REGION Network 8: FT-2011: R-201 Tank Flow from T-101 Totalizer
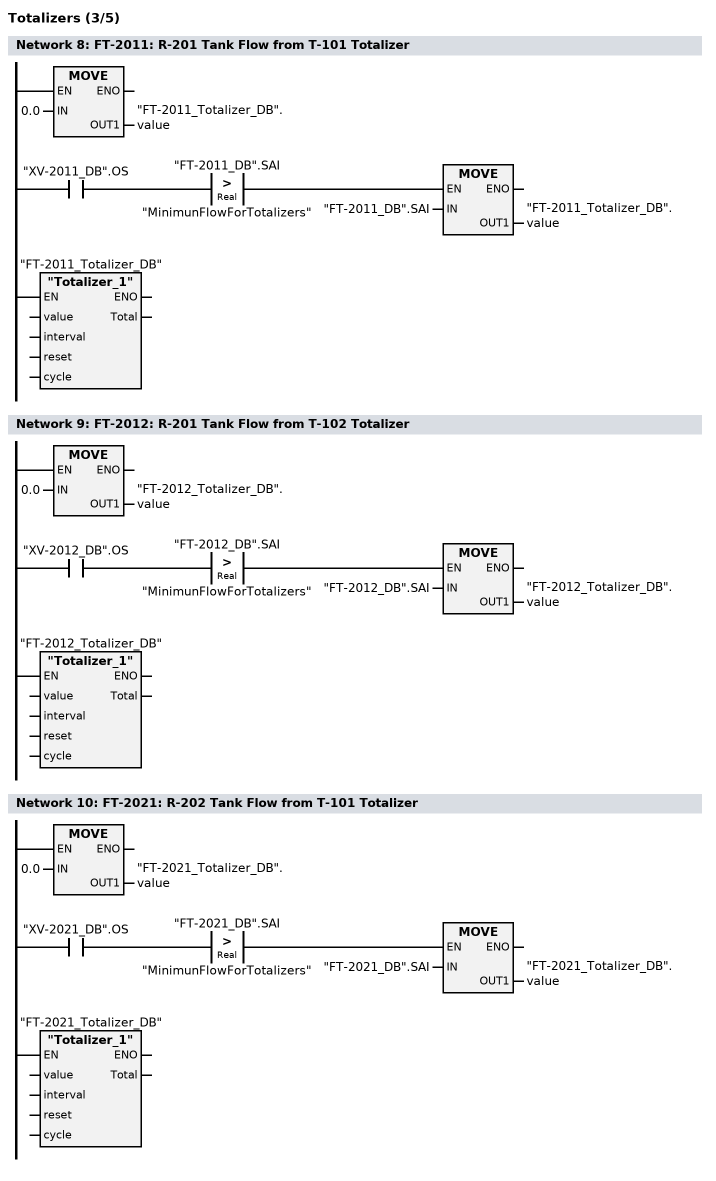
   RUNG wire#powerrail
      { S7_GenerateENO := "TRUE" } Move(in := 0.0, out1 => "FT-2011_Totalizer_DB".value)
   END_RUNG
   RUNG wire#powerrail
      Contact( "XV-2011_DB".OS )
      { S7_Templates := "SrcType := Real" } GT_Contact(in1 := "FT-2011_DB".SAI, in2 := "MinimunFlowForTotalizers")
      { S7_GenerateENO := "TRUE" } Move(in := "FT-2011_DB".SAI, out1 => "FT-2011_Totalizer_DB".value)
   END_RUNG
   RUNG wire#powerrail
      "FT-2011_Totalizer_DB"(value :=, interval :=, reset :=, cycle :=, Total =>)
   END_RUNG
   // the same network as SCL:
   "FT-2011_Totalizer_DB".value := 0.0;
   IF "XV-2011_DB".OS AND ("FT-2011_DB".SAI > "MinimunFlowForTotalizers") THEN
       "FT-2011_Totalizer_DB".value := "FT-2011_DB".SAI;
   END_IF;
   "FT-2011_Totalizer_DB"();   // "Totalizer_1"
END_REGION

REGION Network 9: FT-2012: R-201 Tank Flow from T-102 Totalizer
   RUNG wire#powerrail
      { S7_GenerateENO := "TRUE" } Move(in := 0.0, out1 => "FT-2012_Totalizer_DB".value)
   END_RUNG
   RUNG wire#powerrail
      Contact( "XV-2012_DB".OS )
      { S7_Templates := "SrcType := Real" } GT_Contact(in1 := "FT-2012_DB".SAI, in2 := "MinimunFlowForTotalizers")
      { S7_GenerateENO := "TRUE" } Move(in := "FT-2012_DB".SAI, out1 => "FT-2012_Totalizer_DB".value)
   END_RUNG
   RUNG wire#powerrail
      "FT-2012_Totalizer_DB"(value :=, interval :=, reset :=, cycle :=, Total =>)
   END_RUNG
   // the same network as SCL:
   "FT-2012_Totalizer_DB".value := 0.0;
   IF "XV-2012_DB".OS AND ("FT-2012_DB".SAI > "MinimunFlowForTotalizers") THEN
       "FT-2012_Totalizer_DB".value := "FT-2012_DB".SAI;
   END_IF;
   "FT-2012_Totalizer_DB"();   // "Totalizer_1"
END_REGION

REGION Network 10: FT-2021: R-202 Tank Flow from T-101 Totalizer
   RUNG wire#powerrail
      { S7_GenerateENO := "TRUE" } Move(in := 0.0, out1 => "FT-2021_Totalizer_DB".value)
   END_RUNG
   RUNG wire#powerrail
      Contact( "XV-2021_DB".OS )
      { S7_Templates := "SrcType := Real" } GT_Contact(in1 := "FT-2021_DB".SAI, in2 := "MinimunFlowForTotalizers")
      { S7_GenerateENO := "TRUE" } Move(in := "FT-2021_DB".SAI, out1 => "FT-2021_Totalizer_DB".value)
   END_RUNG
   RUNG wire#powerrail
      "FT-2021_Totalizer_DB"(value :=, interval :=, reset :=, cycle :=, Total =>)
   END_RUNG
   // the same network as SCL:
   "FT-2021_Totalizer_DB".value := 0.0;
   IF "XV-2021_DB".OS AND ("FT-2021_DB".SAI > "MinimunFlowForTotalizers") THEN
       "FT-2021_Totalizer_DB".value := "FT-2021_DB".SAI;
   END_IF;
   "FT-2021_Totalizer_DB"();   // "Totalizer_1"
END_REGION

REGION Network 11: test
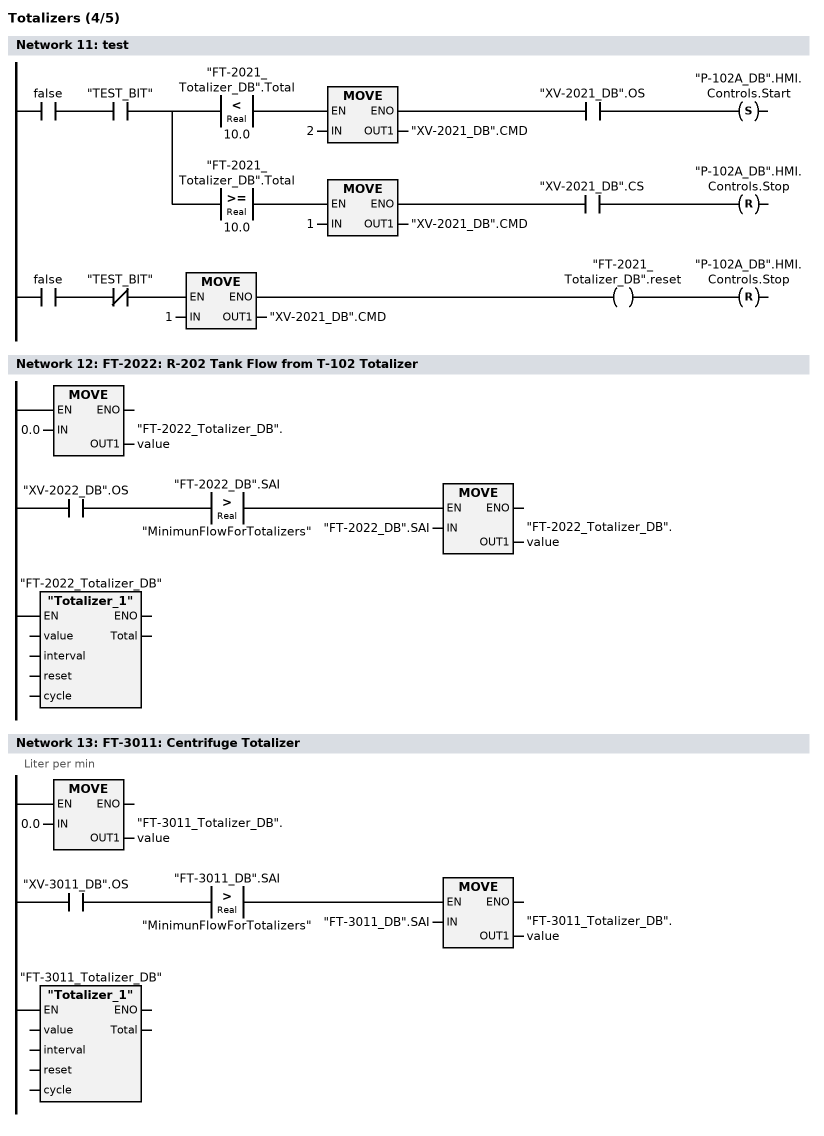
   RUNG wire#powerrail
      Contact( false )
      Contact( "TEST_BIT" )
      wire#w1
      { S7_Templates := "SrcType := Real" } LT_Contact(in1 := "FT-2021_Totalizer_DB".Total, in2 := 10.0)
      { S7_GenerateENO := "TRUE" } Move(in := 2, out1 => "XV-2021_DB".CMD)
      Contact( "XV-2021_DB".OS )
      S_Coil( "P-102A_DB".HMI.Controls.Start )
   END_RUNG
   RUNG wire#w1
      { S7_Templates := "SrcType := Real" } GE_Contact(in1 := "FT-2021_Totalizer_DB".Total, in2 := 10.0)
      { S7_GenerateENO := "TRUE" } Move(in := 1, out1 => "XV-2021_DB".CMD)
      Contact( "XV-2021_DB".CS )
      R_Coil( "P-102A_DB".HMI.Controls.Stop )
   END_RUNG
   RUNG wire#powerrail
      Contact( false )
      I_Contact( "TEST_BIT" )
      { S7_GenerateENO := "TRUE" } Move(in := 1, out1 => "XV-2021_DB".CMD)
      Coil( "FT-2021_Totalizer_DB".reset )
      R_Coil( "P-102A_DB".HMI.Controls.Stop )
   END_RUNG
   // the same network as SCL:
   // ENO of a box is taken as its EN; it also drops when the box reports an error
   #_w1 := false AND "TEST_BIT";
   #_w2 := #_w1 AND ("FT-2021_Totalizer_DB".Total < 10.0);
   IF #_w2 THEN "XV-2021_DB".CMD := 2; END_IF;
   IF #_w2 AND "XV-2021_DB".OS THEN "P-102A_DB".HMI.Controls.Start := TRUE; END_IF;
   #_w3 := #_w1 AND ("FT-2021_Totalizer_DB".Total >= 10.0);
   IF #_w3 THEN "XV-2021_DB".CMD := 1; END_IF;
   IF #_w3 AND "XV-2021_DB".CS THEN "P-102A_DB".HMI.Controls.Stop := FALSE; END_IF;
   #_w4 := false AND NOT "TEST_BIT";
   IF #_w4 THEN "XV-2021_DB".CMD := 1; END_IF;
   "FT-2021_Totalizer_DB".reset := #_w4;
   IF #_w4 THEN "P-102A_DB".HMI.Controls.Stop := FALSE; END_IF;
END_REGION

REGION Network 12: FT-2022: R-202 Tank Flow from T-102 Totalizer
   RUNG wire#powerrail
      { S7_GenerateENO := "TRUE" } Move(in := 0.0, out1 => "FT-2022_Totalizer_DB".value)
   END_RUNG
   RUNG wire#powerrail
      Contact( "XV-2022_DB".OS )
      { S7_Templates := "SrcType := Real" } GT_Contact(in1 := "FT-2022_DB".SAI, in2 := "MinimunFlowForTotalizers")
      { S7_GenerateENO := "TRUE" } Move(in := "FT-2022_DB".SAI, out1 => "FT-2022_Totalizer_DB".value)
   END_RUNG
   RUNG wire#powerrail
      "FT-2022_Totalizer_DB"(value :=, interval :=, reset :=, cycle :=, Total =>)
   END_RUNG
   // the same network as SCL:
   "FT-2022_Totalizer_DB".value := 0.0;
   IF "XV-2022_DB".OS AND ("FT-2022_DB".SAI > "MinimunFlowForTotalizers") THEN
       "FT-2022_Totalizer_DB".value := "FT-2022_DB".SAI;
   END_IF;
   "FT-2022_Totalizer_DB"();   // "Totalizer_1"
END_REGION

REGION Network 13: FT-3011: Centrifuge Totalizer
   // Liter per min
   RUNG wire#powerrail
      { S7_GenerateENO := "TRUE" } Move(in := 0.0, out1 => "FT-3011_Totalizer_DB".value)
   END_RUNG
   RUNG wire#powerrail
      Contact( "XV-3011_DB".OS )
      { S7_Templates := "SrcType := Real" } GT_Contact(in1 := "FT-3011_DB".SAI, in2 := "MinimunFlowForTotalizers")
      { S7_GenerateENO := "TRUE" } Move(in := "FT-3011_DB".SAI, out1 => "FT-3011_Totalizer_DB".value)
   END_RUNG
   RUNG wire#powerrail
      "FT-3011_Totalizer_DB"(value :=, interval :=, reset :=, cycle :=, Total =>)
   END_RUNG
   // the same network as SCL:
   "FT-3011_Totalizer_DB".value := 0.0;
   IF "XV-3011_DB".OS AND ("FT-3011_DB".SAI > "MinimunFlowForTotalizers") THEN
       "FT-3011_Totalizer_DB".value := "FT-3011_DB".SAI;
   END_IF;
   "FT-3011_Totalizer_DB"();   // "Totalizer_1"
END_REGION

REGION Network 14: FT-3012:Centrifuge Dry Spin Totalizer
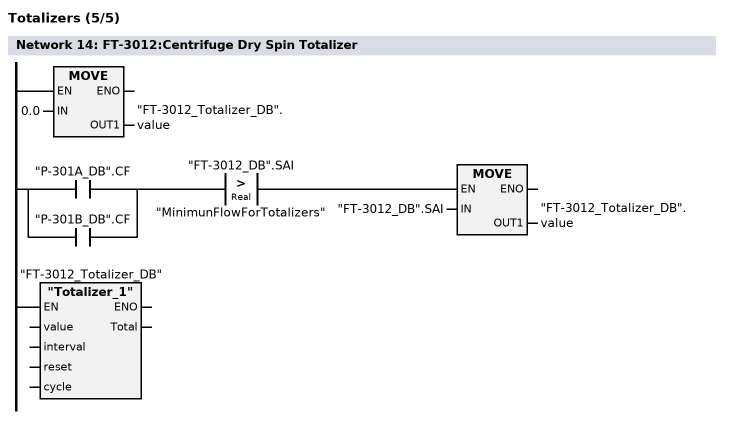
   RUNG wire#powerrail
      { S7_GenerateENO := "TRUE" } Move(in := 0.0, out1 => "FT-3012_Totalizer_DB".value)
   END_RUNG
   RUNG wire#powerrail
      Contact( "P-301A_DB".CF )
      wire#w1
      { S7_Templates := "SrcType := Real" } GT_Contact(in1 := "FT-3012_DB".SAI, in2 := "MinimunFlowForTotalizers")
      { S7_GenerateENO := "TRUE" } Move(in := "FT-3012_DB".SAI, out1 => "FT-3012_Totalizer_DB".value)
   END_RUNG
   RUNG wire#powerrail
      Contact( "P-301B_DB".CF )
   END_RUNG wire#w1
   RUNG wire#powerrail
      "FT-3012_Totalizer_DB"(value :=, interval :=, reset :=, cycle :=, Total =>)
   END_RUNG
   // the same network as SCL:
   "FT-3012_Totalizer_DB".value := 0.0;
   IF ("P-301A_DB".CF OR "P-301B_DB".CF) AND ("FT-3012_DB".SAI > "MinimunFlowForTotalizers") THEN
       "FT-3012_Totalizer_DB".value := "FT-3012_DB".SAI;
   END_IF;
   "FT-3012_Totalizer_DB"();   // "Totalizer_1"
END_REGION
END_FUNCTION

// folder: VFD

FUNCTION "VFD" : Void   // FC25, LAD
{ S7_Optimized_Access := 'TRUE' }
VERSION : 0.1
   VAR_TEMP
      "T-101" : Real;
      "T-102" : Real;
   END_VAR
BEGIN

REGION Network 1: VFD-1011A: Tank T-101 Agitator
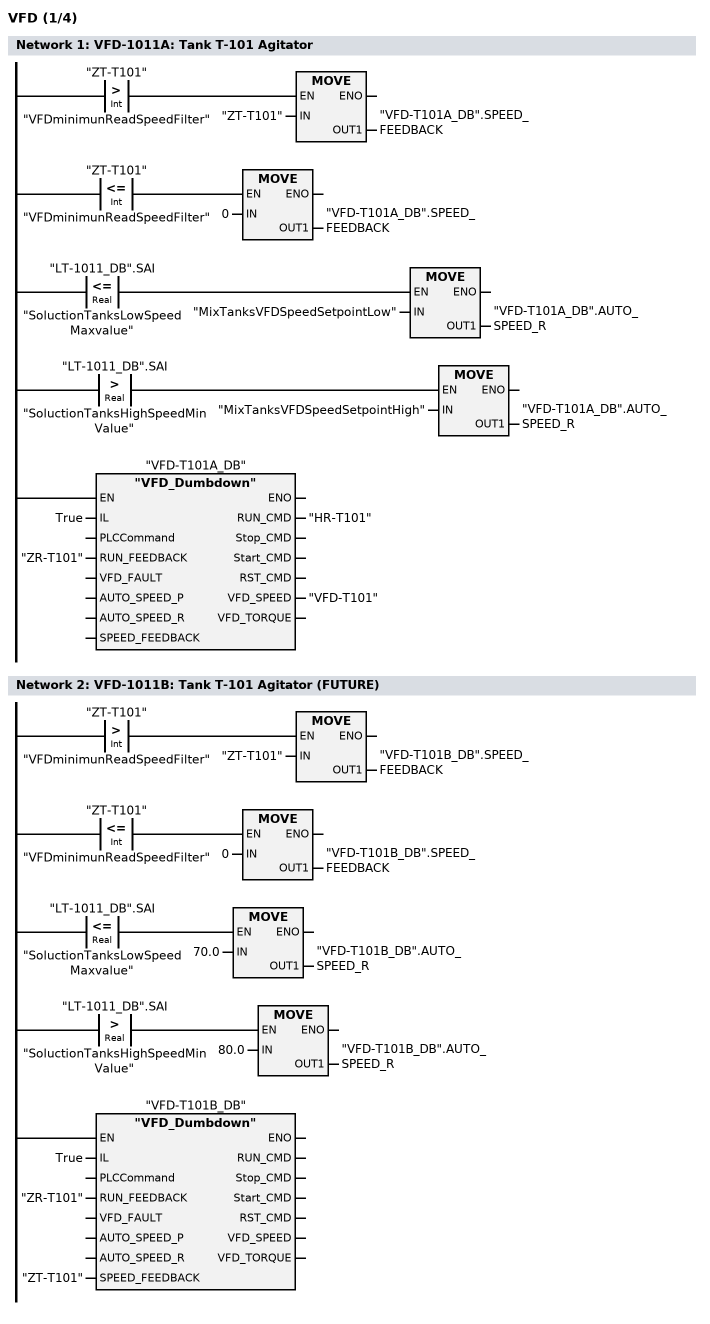
   RUNG wire#powerrail
      { S7_Templates := "SrcType := Int" } GT_Contact(in1 := "ZT-T101", in2 := "VFDminimunReadSpeedFilter")
      { S7_GenerateENO := "TRUE" } Move(in := "ZT-T101", out1 => "VFD-T101A_DB".SPEED_FEEDBACK)
   END_RUNG
   RUNG wire#powerrail
      { S7_Templates := "SrcType := Int" } LE_Contact(in1 := "ZT-T101", in2 := "VFDminimunReadSpeedFilter")
      { S7_GenerateENO := "TRUE" } Move(in := 0, out1 => "VFD-T101A_DB".SPEED_FEEDBACK)
   END_RUNG
   RUNG wire#powerrail
      { S7_Templates := "SrcType := Real" } LE_Contact(in1 := "LT-1011_DB".SAI, in2 := "SoluctionTanksLowSpeedMaxvalue")
      { S7_GenerateENO := "TRUE" } Move(in := "MixTanksVFDSpeedSetpointLow", out1 => "VFD-T101A_DB".AUTO_SPEED_R)
   END_RUNG
   RUNG wire#powerrail
      { S7_Templates := "SrcType := Real" } GT_Contact(in1 := "LT-1011_DB".SAI, in2 := "SoluctionTanksHighSpeedMinValue")
      { S7_GenerateENO := "TRUE" } Move(in := "MixTanksVFDSpeedSetpointHigh", out1 => "VFD-T101A_DB".AUTO_SPEED_R)
   END_RUNG
   RUNG wire#powerrail
      "VFD-T101A_DB"(IL := True, PLCCommand :=, RUN_FEEDBACK := "ZR-T101", VFD_FAULT :=, AUTO_SPEED_P :=, AUTO_SPEED_R :=, SPEED_FEEDBACK :=, RUN_CMD => "HR-T101", Stop_CMD =>, Start_CMD =>, RST_CMD =>, VFD_SPEED => "VFD-T101", VFD_TORQUE =>)
   END_RUNG
   // the same network as SCL:
   IF "ZT-T101" > "VFDminimunReadSpeedFilter" THEN "VFD-T101A_DB".SPEED_FEEDBACK := "ZT-T101"; END_IF;
   IF "ZT-T101" <= "VFDminimunReadSpeedFilter" THEN "VFD-T101A_DB".SPEED_FEEDBACK := 0; END_IF;
   IF "LT-1011_DB".SAI <= "SoluctionTanksLowSpeedMaxvalue" THEN
       "VFD-T101A_DB".AUTO_SPEED_R := "MixTanksVFDSpeedSetpointLow";
   END_IF;
   IF "LT-1011_DB".SAI > "SoluctionTanksHighSpeedMinValue" THEN
       "VFD-T101A_DB".AUTO_SPEED_R := "MixTanksVFDSpeedSetpointHigh";
   END_IF;
   "VFD-T101A_DB"(IL := True, RUN_FEEDBACK := "ZR-T101", RUN_CMD => "HR-T101", VFD_SPEED => "VFD-T101");   // "VFD_Dumbdown"
END_REGION

REGION Network 2: VFD-1011B: Tank T-101 Agitator (FUTURE)
   RUNG wire#powerrail
      { S7_Templates := "SrcType := Int" } GT_Contact(in1 := "ZT-T101", in2 := "VFDminimunReadSpeedFilter")
      { S7_GenerateENO := "TRUE" } Move(in := "ZT-T101", out1 => "VFD-T101B_DB".SPEED_FEEDBACK)
   END_RUNG
   RUNG wire#powerrail
      { S7_Templates := "SrcType := Int" } LE_Contact(in1 := "ZT-T101", in2 := "VFDminimunReadSpeedFilter")
      { S7_GenerateENO := "TRUE" } Move(in := 0, out1 => "VFD-T101B_DB".SPEED_FEEDBACK)
   END_RUNG
   RUNG wire#powerrail
      { S7_Templates := "SrcType := Real" } LE_Contact(in1 := "LT-1011_DB".SAI, in2 := "SoluctionTanksLowSpeedMaxvalue")
      { S7_GenerateENO := "TRUE" } Move(in := 70.0, out1 => "VFD-T101B_DB".AUTO_SPEED_R)
   END_RUNG
   RUNG wire#powerrail
      { S7_Templates := "SrcType := Real" } GT_Contact(in1 := "LT-1011_DB".SAI, in2 := "SoluctionTanksHighSpeedMinValue")
      { S7_GenerateENO := "TRUE" } Move(in := 80.0, out1 => "VFD-T101B_DB".AUTO_SPEED_R)
   END_RUNG
   RUNG wire#powerrail
      "VFD-T101B_DB"(IL := True, PLCCommand :=, RUN_FEEDBACK := "ZR-T101", VFD_FAULT :=, AUTO_SPEED_P :=, AUTO_SPEED_R :=, SPEED_FEEDBACK := "ZT-T101", RUN_CMD =>, Stop_CMD =>, Start_CMD =>, RST_CMD =>, VFD_SPEED =>, VFD_TORQUE =>)
   END_RUNG
   // the same network as SCL:
   IF "ZT-T101" > "VFDminimunReadSpeedFilter" THEN "VFD-T101B_DB".SPEED_FEEDBACK := "ZT-T101"; END_IF;
   IF "ZT-T101" <= "VFDminimunReadSpeedFilter" THEN "VFD-T101B_DB".SPEED_FEEDBACK := 0; END_IF;
   IF "LT-1011_DB".SAI <= "SoluctionTanksLowSpeedMaxvalue" THEN "VFD-T101B_DB".AUTO_SPEED_R := 70.0; END_IF;
   IF "LT-1011_DB".SAI > "SoluctionTanksHighSpeedMinValue" THEN "VFD-T101B_DB".AUTO_SPEED_R := 80.0; END_IF;
   "VFD-T101B_DB"(IL := True, RUN_FEEDBACK := "ZR-T101", SPEED_FEEDBACK := "ZT-T101");   // "VFD_Dumbdown"
END_REGION

REGION Network 3: VFD-1021A: Tank T-102 Agitator
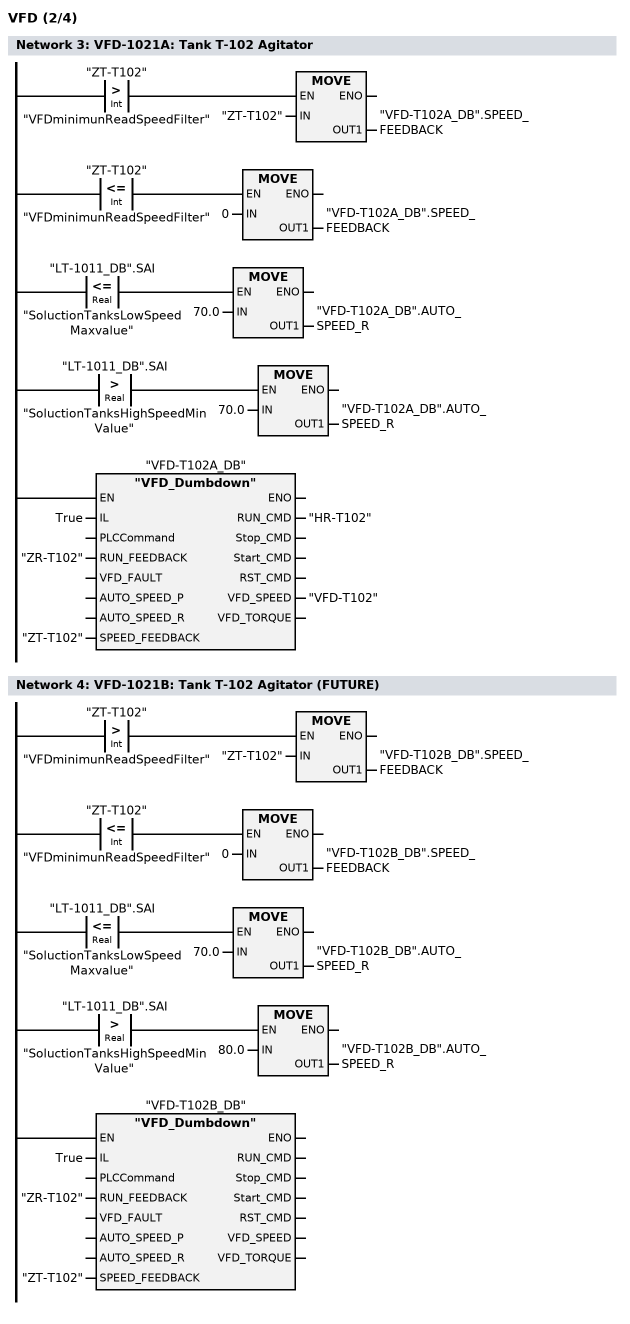
   RUNG wire#powerrail
      { S7_Templates := "SrcType := Int" } GT_Contact(in1 := "ZT-T102", in2 := "VFDminimunReadSpeedFilter")
      { S7_GenerateENO := "TRUE" } Move(in := "ZT-T102", out1 => "VFD-T102A_DB".SPEED_FEEDBACK)
   END_RUNG
   RUNG wire#powerrail
      { S7_Templates := "SrcType := Int" } LE_Contact(in1 := "ZT-T102", in2 := "VFDminimunReadSpeedFilter")
      { S7_GenerateENO := "TRUE" } Move(in := 0, out1 => "VFD-T102A_DB".SPEED_FEEDBACK)
   END_RUNG
   RUNG wire#powerrail
      { S7_Templates := "SrcType := Real" } LE_Contact(in1 := "LT-1011_DB".SAI, in2 := "SoluctionTanksLowSpeedMaxvalue")
      { S7_GenerateENO := "TRUE" } Move(in := 70.0, out1 => "VFD-T102A_DB".AUTO_SPEED_R)
   END_RUNG
   RUNG wire#powerrail
      { S7_Templates := "SrcType := Real" } GT_Contact(in1 := "LT-1011_DB".SAI, in2 := "SoluctionTanksHighSpeedMinValue")
      { S7_GenerateENO := "TRUE" } Move(in := 70.0, out1 => "VFD-T102A_DB".AUTO_SPEED_R)
   END_RUNG
   RUNG wire#powerrail
      "VFD-T102A_DB"(IL := True, PLCCommand :=, RUN_FEEDBACK := "ZR-T102", VFD_FAULT :=, AUTO_SPEED_P :=, AUTO_SPEED_R :=, SPEED_FEEDBACK := "ZT-T102", RUN_CMD => "HR-T102", Stop_CMD =>, Start_CMD =>, RST_CMD =>, VFD_SPEED => "VFD-T102", VFD_TORQUE =>)
   END_RUNG
   // the same network as SCL:
   IF "ZT-T102" > "VFDminimunReadSpeedFilter" THEN "VFD-T102A_DB".SPEED_FEEDBACK := "ZT-T102"; END_IF;
   IF "ZT-T102" <= "VFDminimunReadSpeedFilter" THEN "VFD-T102A_DB".SPEED_FEEDBACK := 0; END_IF;
   IF "LT-1011_DB".SAI <= "SoluctionTanksLowSpeedMaxvalue" THEN "VFD-T102A_DB".AUTO_SPEED_R := 70.0; END_IF;
   IF "LT-1011_DB".SAI > "SoluctionTanksHighSpeedMinValue" THEN "VFD-T102A_DB".AUTO_SPEED_R := 70.0; END_IF;
   "VFD-T102A_DB"(IL := True,   // "VFD_Dumbdown"
                  RUN_FEEDBACK := "ZR-T102",
                  SPEED_FEEDBACK := "ZT-T102",
                  RUN_CMD => "HR-T102",
                  VFD_SPEED => "VFD-T102");
END_REGION

REGION Network 4: VFD-1021B: Tank T-102 Agitator (FUTURE)
   RUNG wire#powerrail
      { S7_Templates := "SrcType := Int" } GT_Contact(in1 := "ZT-T102", in2 := "VFDminimunReadSpeedFilter")
      { S7_GenerateENO := "TRUE" } Move(in := "ZT-T102", out1 => "VFD-T102B_DB".SPEED_FEEDBACK)
   END_RUNG
   RUNG wire#powerrail
      { S7_Templates := "SrcType := Int" } LE_Contact(in1 := "ZT-T102", in2 := "VFDminimunReadSpeedFilter")
      { S7_GenerateENO := "TRUE" } Move(in := 0, out1 => "VFD-T102B_DB".SPEED_FEEDBACK)
   END_RUNG
   RUNG wire#powerrail
      { S7_Templates := "SrcType := Real" } LE_Contact(in1 := "LT-1011_DB".SAI, in2 := "SoluctionTanksLowSpeedMaxvalue")
      { S7_GenerateENO := "TRUE" } Move(in := 70.0, out1 => "VFD-T102B_DB".AUTO_SPEED_R)
   END_RUNG
   RUNG wire#powerrail
      { S7_Templates := "SrcType := Real" } GT_Contact(in1 := "LT-1011_DB".SAI, in2 := "SoluctionTanksHighSpeedMinValue")
      { S7_GenerateENO := "TRUE" } Move(in := 80.0, out1 => "VFD-T102B_DB".AUTO_SPEED_R)
   END_RUNG
   RUNG wire#powerrail
      "VFD-T102B_DB"(IL := True, PLCCommand :=, RUN_FEEDBACK := "ZR-T102", VFD_FAULT :=, AUTO_SPEED_P :=, AUTO_SPEED_R :=, SPEED_FEEDBACK := "ZT-T102", RUN_CMD =>, Stop_CMD =>, Start_CMD =>, RST_CMD =>, VFD_SPEED =>, VFD_TORQUE =>)
   END_RUNG
   // the same network as SCL:
   IF "ZT-T102" > "VFDminimunReadSpeedFilter" THEN "VFD-T102B_DB".SPEED_FEEDBACK := "ZT-T102"; END_IF;
   IF "ZT-T102" <= "VFDminimunReadSpeedFilter" THEN "VFD-T102B_DB".SPEED_FEEDBACK := 0; END_IF;
   IF "LT-1011_DB".SAI <= "SoluctionTanksLowSpeedMaxvalue" THEN "VFD-T102B_DB".AUTO_SPEED_R := 70.0; END_IF;
   IF "LT-1011_DB".SAI > "SoluctionTanksHighSpeedMinValue" THEN "VFD-T102B_DB".AUTO_SPEED_R := 80.0; END_IF;
   "VFD-T102B_DB"(IL := True, RUN_FEEDBACK := "ZR-T102", SPEED_FEEDBACK := "ZT-T102");   // "VFD_Dumbdown"
END_REGION

REGION Network 5: VFD-1031: Tank T-103 Agitator (FUTURE)
   // "ZR-C301R"
   // "ZT-R201"
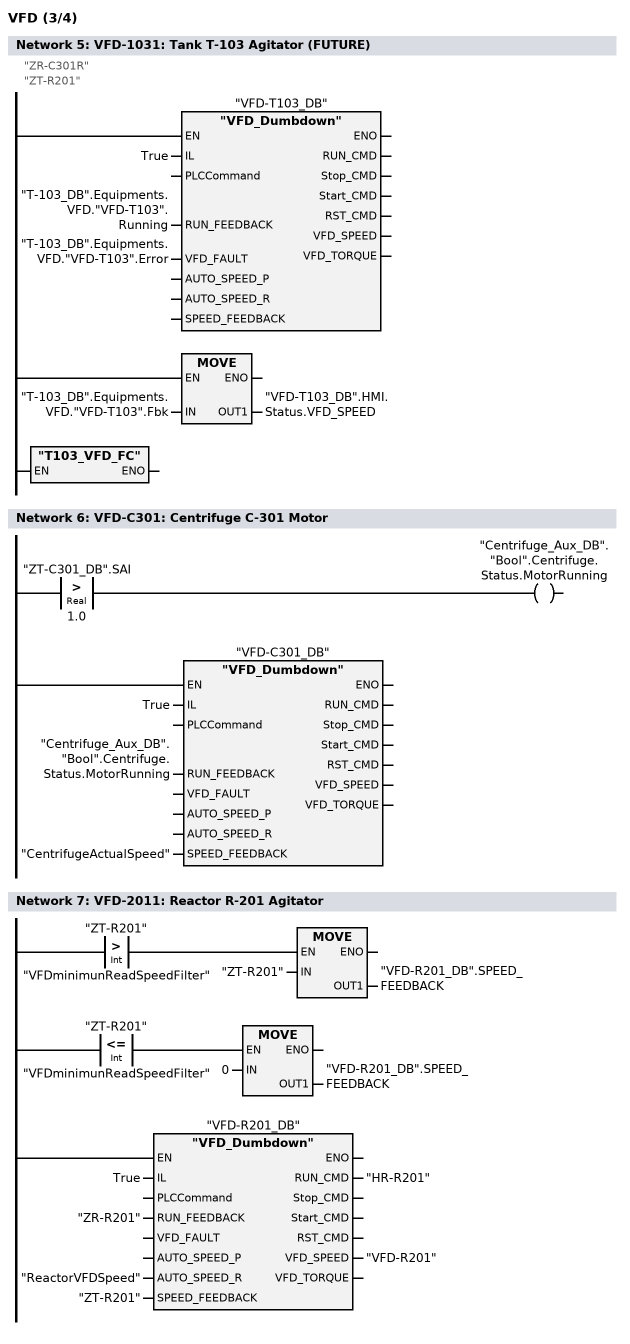
   RUNG wire#powerrail
      "VFD-T103_DB"(IL := True, PLCCommand :=, RUN_FEEDBACK := "T-103_DB".Equipments.VFD."VFD-T103".Running, VFD_FAULT := "T-103_DB".Equipments.VFD."VFD-T103".Error, AUTO_SPEED_P :=, AUTO_SPEED_R :=, SPEED_FEEDBACK :=, RUN_CMD =>, Stop_CMD =>, Start_CMD =>, RST_CMD =>, VFD_SPEED =>, VFD_TORQUE =>)
   END_RUNG
   RUNG wire#powerrail
      Move(in := "T-103_DB".Equipments.VFD."VFD-T103".Fbk, out1 => "VFD-T103_DB".HMI.Status.VFD_SPEED)
   END_RUNG
   RUNG wire#powerrail
      "T103_VFD_FC"()
   END_RUNG
   // the same network as SCL:
   "VFD-T103_DB"(IL := True,   // "VFD_Dumbdown"
                 RUN_FEEDBACK := "T-103_DB".Equipments.VFD."VFD-T103".Running,
                 VFD_FAULT := "T-103_DB".Equipments.VFD."VFD-T103".Error);
   "VFD-T103_DB".HMI.Status.VFD_SPEED := "T-103_DB".Equipments.VFD."VFD-T103".Fbk;
   "T103_VFD_FC"();
END_REGION

REGION Network 6: VFD-C301: Centrifuge C-301 Motor
   RUNG wire#powerrail
      { S7_Templates := "SrcType := Real" } GT_Contact(in1 := "ZT-C301_DB".SAI, in2 := 1.0)
      Coil( "Centrifuge_Aux_DB"."Bool".Centrifuge.Status.MotorRunning )
   END_RUNG
   RUNG wire#powerrail
      "VFD-C301_DB"(IL := True, PLCCommand :=, RUN_FEEDBACK := "Centrifuge_Aux_DB"."Bool".Centrifuge.Status.MotorRunning, VFD_FAULT :=, AUTO_SPEED_P :=, AUTO_SPEED_R :=, SPEED_FEEDBACK := "CentrifugeActualSpeed", RUN_CMD =>, Stop_CMD =>, Start_CMD =>, RST_CMD =>, VFD_SPEED =>, VFD_TORQUE =>)
   END_RUNG
   // the same network as SCL:
   "Centrifuge_Aux_DB"."Bool".Centrifuge.Status.MotorRunning := "ZT-C301_DB".SAI > 1.0;
   "VFD-C301_DB"(IL := True,   // "VFD_Dumbdown"
                 RUN_FEEDBACK := "Centrifuge_Aux_DB"."Bool".Centrifuge.Status.MotorRunning,
                 SPEED_FEEDBACK := "CentrifugeActualSpeed");
END_REGION

REGION Network 7: VFD-2011: Reactor R-201 Agitator
   RUNG wire#powerrail
      { S7_Templates := "SrcType := Int" } GT_Contact(in1 := "ZT-R201", in2 := "VFDminimunReadSpeedFilter")
      { S7_GenerateENO := "TRUE" } Move(in := "ZT-R201", out1 => "VFD-R201_DB".SPEED_FEEDBACK)
   END_RUNG
   RUNG wire#powerrail
      { S7_Templates := "SrcType := Int" } LE_Contact(in1 := "ZT-R201", in2 := "VFDminimunReadSpeedFilter")
      { S7_GenerateENO := "TRUE" } Move(in := 0, out1 => "VFD-R201_DB".SPEED_FEEDBACK)
   END_RUNG
   RUNG wire#powerrail
      "VFD-R201_DB"(IL := True, PLCCommand :=, RUN_FEEDBACK := "ZR-R201", VFD_FAULT :=, AUTO_SPEED_P :=, AUTO_SPEED_R := "ReactorVFDSpeed", SPEED_FEEDBACK := "ZT-R201", RUN_CMD => "HR-R201", Stop_CMD =>, Start_CMD =>, RST_CMD =>, VFD_SPEED => "VFD-R201", VFD_TORQUE =>)
   END_RUNG
   // the same network as SCL:
   IF "ZT-R201" > "VFDminimunReadSpeedFilter" THEN "VFD-R201_DB".SPEED_FEEDBACK := "ZT-R201"; END_IF;
   IF "ZT-R201" <= "VFDminimunReadSpeedFilter" THEN "VFD-R201_DB".SPEED_FEEDBACK := 0; END_IF;
   "VFD-R201_DB"(IL := True,   // "VFD_Dumbdown"
                 RUN_FEEDBACK := "ZR-R201",
                 AUTO_SPEED_R := "ReactorVFDSpeed",
                 SPEED_FEEDBACK := "ZT-R201",
                 RUN_CMD => "HR-R201",
                 VFD_SPEED => "VFD-R201");
END_REGION

REGION Network 8: "VFD-2021: Reactor R-202 Agitator